(* Logix 5000 project; controller PLC_MCC1300_75F1 vendor 1 type 14 code 166 rev 32.11; software revision 32.04; part 65 of 83 *)
(* tags used below, declared in another part *)
   CM_AreaStackerToLine_JS1 : CM_AreaStackerToLine;
   CM_AreaStackerToLine_JS1_Sync : CM_AreaStackerToLine;
   CONST_dDest_Cullet : DINT;
   CONST_dDest_Stk : DINT;
   CONST_rgdDestMask : DINT[32];   // Destination Mask
   Convoy_SL_DATA_NULL : UDT_Convoy_SL;
   GP_AccessArea_M316S_STC : GP_AccessArea_STC;
   GP_CheckIdPlatePresent : GP_CheckIdPlatePresent;
   GP_InvertCapxLite : GP_InvertCapxLite;
   GP_M316A : GP_Rotator;
   GP_OB_InitializeMain : GP_OB_Initialize;
   GP_RampSpace : GP_RampSpace;
   Gp_SpaceConvUtilities_V1 : GP_SpaceConvUtilities_V1;
   M310B : MAC_Conveyor;
   M310B_Data : UDT_Convoy_SL;
   M310B_SpaceConv_Utilities : SpaceConv_Utilities;
   M312 : MAC_Conveyor_Single;
   M312_SpaceConv_Utilities : SpaceConv_Utilities;
   M315A_SpaceConv_Utilities : SpaceConv_Utilities;
   M315B : MAC_Conveyor;
   M315B_Data : UDT_Convoy_SL;
   M315B_SpaceConv_Utilities : SpaceConv_Utilities;
   M316 : MAC_Conveyor;
   M316_ALM : MAC_Conveyor_ALM;
   M316_Data : UDT_Convoy_SL;
   M316_dLastRotationA_ID : DINT;
   M316_HMW : MAC_Conveyor_HMW;
   M316_M1_DR_IN_MAM : MOTION_INSTRUCTION;
   M316_SpaceConv_Utilities : SpaceConv_Utilities;
   M316_xOS_SentToCullet : BOOL;
   M316_xPlateCullet : BOOL;
   M316_xSendCulletReqActive : BOOL;
   M316A : MAC_Rotator;
   M316A_Data : UDT_Convoy_SL;
   M316A_HMR : MAC_Rotator_HMR;
   M316A_HMW : MAC_Rotator_HMW;
   M316A_M1_DR : AXIS_CIP_DRIVE;
   M316A_M1_DR_IN_MAM : MOTION_INSTRUCTION;
   M316A_rLastPosition : REAL;
   M317_SpaceConv_Utilities : SpaceConv_Utilities;
   Sbr_OUT_ReqRot_CW : BOOL;
   TMP_d : DINT;
   TMP_dActualOnLHS : DINT;
   TMP_dConveyorNumberForZoneCleaning : DINT;
   TMP_dDecelerationPositionEndConveyor : DINT;
   TMP_dMissingOnLHS : DINT;
   TMP_dOffsetLoadUnload_cmm : DINT;
   TMP_dPhEndPosition_cmm : DINT;
   TMP_HeadPos : DINT;
   TMP_Portrait : BOOL;
   TMP_rgxId : DINT[10];
   TMP_x : BOOL;
   TMP_xConveyorInvolvedInCleaning : BOOL;
   TMP_xConveyorOfStartCleaning : BOOL;
   TMP_xCulletPresent : BOOL;
   TMP_xEnableLoadUnload : BOOL;
   TMP_xEnableZoneCleaning : BOOL;
   TMP_xJustOnePlateMissing : BOOL;
   TMP_xLiteThisDestPresent : BOOL;
   x316PortraitMode : BOOL;
   xAlwaysOFF : BOOL;
   xAlwaysON : BOOL;
   xDebugOFF : BOOL;
   Z402 : MAC_Zone;
   Z402_HMR : MAC_Zone_HMR;
   Z402_HMW : MAC_Zone_HMW;
(* MainProgram, continued *)

ROUTINE M316_Alarm   (* ladder *)
   // Reset Alarm
   0: XIC(Z402.tmON_ResetAlarm.DN)FLL(0,M316_ALM,1);
   1: XIC(Z402.ST_xEnableControlError)XIC(M316.INPUT_xDriveError_M1)OTL(M316_ALM.rgxStoppingFault_M[0].1);
   2: XIC(Z402.ST_xEnableControlError)XIO(M316.INPUT_xDriveError_M1)[XIC(M316.OUTPUT_xRun_M1) ,XIC(M316.OUTPUT_xReverse_M1) ,XIC(M316.OUTPUT_xPositioning_M1) ]XIO(M316.INPUT_xDriveFeedback_M1)[XIO(M316.tmON_FeedbackTimeOut_M1.DN) TON(M316.tmON_FeedbackTimeOut_M1,?,?) ,XIC(M316.tmON_FeedbackTimeOut_M1.DN) OTL(M316_ALM.rgxStoppingFault_M[0].2) ];
   3: XIC(Z402.ST_xEnableControlError)XIO(M316.INPUT_xMotorThermalProbe_M1)OTL(M316_ALM.rgxStoppingFault_M[0].4);
   4: XIC(Z402.ST_xEnableControlError)[XIC(M316.INPUT_xDriveInhibit_M1) ,XIC(M316.OUTPUT_xDriveEnable_M1) XIO(M316.INPUT_xDriveReady_M1) ][XIO(M316.tmON_DriveInhibit_M1.DN) TON(M316.tmON_DriveInhibit_M1,?,?) ,XIC(M316.tmON_DriveInhibit_M1.DN) OTL(M316_ALM.rgxStoppingFault_M[0].6) ];
   5: XIC(Z402.ST_xEnableControlError)XIC(M316.INPUT_xDriveError_M2)OTL(M316_ALM.rgxStoppingFault_M[0].11);
   6: XIC(Z402.ST_xEnableControlError)XIO(M316.INPUT_xDriveError_M2)[XIC(M316.OUTPUT_xRun_M2) ,XIC(M316.OUTPUT_xReverse_M2) ,XIC(M316.OUTPUT_xPositioning_M2) ]XIO(M316.INPUT_xDriveFeedback_M2)[XIO(M316.tmON_FeedbackTimeOut_M2.DN) TON(M316.tmON_FeedbackTimeOut_M2,?,?) ,XIC(M316.tmON_FeedbackTimeOut_M2.DN) OTL(M316_ALM.rgxStoppingFault_M[0].12) ];
   7: XIC(Z402.ST_xEnableControlError)XIO(M316.INPUT_xMotorThermalProbe_M2)OTL(M316_ALM.rgxStoppingFault_M[0].14);
   8: XIC(Z402.ST_xEnableControlError)[XIC(M316.INPUT_xDriveInhibit_M2) ,XIC(M316.OUTPUT_xDriveEnable_M2) XIO(M316.INPUT_xDriveReady_M2) ][XIO(M316.tmON_DriveInhibit_M2.DN) TON(M316.tmON_DriveInhibit_M2,?,?) ,XIC(M316.tmON_DriveInhibit_M2.DN) OTL(M316_ALM.rgxStoppingFault_M[0].16) ];
   9: XIC(M316.ST_xEnableControlError)XIC(M316.PH_x.7)NEQ(M316_SpaceConv_Utilities.CONST_dSyncMode,0)[XIO(M316.ST_xPlateSynchronized) OTL(M316_ALM.rgxWarning[0].0) ,XIC(M316.ST_xPlateSynchronized) OTU(M316_ALM.rgxWarning[0].0) ];
   10: XIC(M316.ST_xEnableControlError)[XIC(M316_Data.tFlag.tConveyor.xReqStop) [XIC(M316.PH_x.0) ,XIC(M316.PH_x.1) ] ADD(M316_SpaceConv_Utilities.CONST_dConveyorLength_cmm,200000,TMP_d) GRT(M316_SpaceConv_Utilities.O_dHeadPosition_cmm,TMP_d) ,XIC(M316.PH_x.16) CPT(TMP_d,M316_SpaceConv_Utilities.CONST_dConveyorLength_cmm + M316.AUX_dDecSpace_cmm) GRT(M316_SpaceConv_Utilities.O_dHeadPosition_cmm,TMP_d) ][OTL(M316_ALM.rgxWarning[0].1) ,OTL(M316.ST_xPhaseError) ];
   11: XIC(M316.ST_xEnableControlError)[XIC(M316.PH_x.0) ,XIC(M316.PH_x.8) ,XIC(M316.PH_x.16) ]XIO(M316A.INPUT_xLowPosition)OTL(M316_ALM.rgxStoppingFault[0].0);
   // #####_CUMULATIVE ALARM_#####
   12: NOP();
   13: [NEQ(M316_ALM.rgxStoppingFault[0],0) ,NEQ(M316_ALM.rgxStoppingFault_M[0],0) ,NEQ(M316_ALM.rgxStoppingFault_M[1],0) ]OTE(M316.ST_xStopMachineFault);
   14: [NEQ(M316_ALM.rgxFault[0],0) ,NEQ(M316_ALM.rgxFault_M[0],0) ,NEQ(M316_ALM.rgxFault_M[1],0) ]OTE(M316.ST_xStopNextCycleFault);
END_ROUTINE

ROUTINE M316_Logic   (* ladder *)
   // #####_COSTANTS_#####
   0: [MOV(4030,TMP_dConveyorNumberForZoneCleaning) MOV(350000,TMP_dOffsetLoadUnload_cmm) MOV(500,M316_SpaceConv_Utilities.CONST_dPresetFeedbackTime_ms) OTL(TMP_xEnableLoadUnload) OTU(TMP_xEnableZoneCleaning) MOV(450000,M316_SpaceConv_Utilities.CONST_dConveyorLength_cmm) MOV(375000,M316_SpaceConv_Utilities.CONST_dConveyorWidth_cmm) SUB(M316_SpaceConv_Utilities.CONST_dConveyorLength_cmm,M316.AUX_dAccSpace_cmm,M316.AUX_dPresetStopLoad_cmm) ADD(M316_SpaceConv_Utilities.CONST_dConveyorLength_cmm,M316.AUX_dDecSpace_cmm,M316.AUX_dPresetStopUnload_cmm) MOV(1.2,M316_SpaceConv_Utilities.CONST_rAcceleration_ms2) MOV(1.2,M316_SpaceConv_Utilities.CONST_rDeceleration_ms2) MOV(M316_SpaceConv_Utilities.CONST_dConveyorLength_cmm,TMP_dPhEndPosition_cmm) ,XIO(M316.PH_x.22) [MOV(1,M316_SpaceConv_Utilities.CONST_dSyncMode) ,MOV(25000,M316_SpaceConv_Utilities.CONST_dSyncroPhPosition_cmm) ,MOV(200000,M316_SpaceConv_Utilities.CONST_dSyncroPhWindow_cmm) ] ,XIC(M316.PH_x.22) [MOV(1,M316_SpaceConv_Utilities.CONST_dSyncMode) ,MOV(0,M316_SpaceConv_Utilities.CONST_dSyncroPhPosition_cmm) ,MOV(300000,M316_SpaceConv_Utilities.CONST_dSyncroPhWindow_cmm) ] ];
   // #####_MATCH_#####
   1: NOP();
   // Conveyor Cleaning
   2: XIC(TMP_xEnableZoneCleaning)XIC(Z402.ST_xCleaningAccepted)GRT(Z402_HMW.dCleaningSelection,0)[EQU(Z402_HMW.dCleaningSelection,TMP_dConveyorNumberForZoneCleaning) OTE(TMP_xConveyorOfStartCleaning) ,GEQ(Z402_HMW.dCleaningSelection,TMP_dConveyorNumberForZoneCleaning) OTE(TMP_xConveyorInvolvedInCleaning) ];
   // Enable control error
   3: XIC(Z402.ST_xEnableControlError)OTE(M316.ST_xEnableControlError);
   // Mode 7 - Offsett for load/unload Simultaney
   4: XIC(M316.PH_x.8)MOV(M316.AUX_dPresetStopLoad_cmm,M316_SpaceConv_Utilities.ST_dStopLoadForseen_cmm)MOV(TMP_dOffsetLoadUnload_cmm,M316_SpaceConv_Utilities.CONF_MD7_dOffset_cmm)GP_SpaceConvUtilities_V1(Gp_SpaceConvUtilities_V1,M316_SpaceConv_Utilities,M315A_SpaceConv_Utilities,M317_SpaceConv_Utilities,7);
   // #####_ALARMS_#####
   5: NOP();
   // Call Alarm Routine
   6: JSR(M316_Alarm,0);
   // Call Alarm Routine
   7: JSR(M316A_Rotator_Alarm,0);
   // #####_HMI_LOGICS_#####
   8: NOP();
   // Condition ok for Cleaning
   9: [XIO(TMP_xEnableZoneCleaning) ,XIC(TMP_xEnableZoneCleaning) XIC(M316.ST_xOutputEnable) [XIO(TMP_xConveyorOfStartCleaning) ,XIC(M316.PH_x.0) ,XIO(M316.PH_x.8) ] ]OTE(M316.ST_xCleaningConditionOK);
   // Cleaning Accepted
   10: [[XIC(M316_HMW.xStopLocalCleaningRequest) ,XIC(Z402_HMW.xStopCleanZoneRequest) ] OTU(M316_HMW.xStopLocalCleaningRequest) OTU(M316_HMW.xLocalCleaningRequest) ,[XIC(M316_HMW.xLocalCleaningRequest) ,XIC(xAlwaysOFF) XIC(M316.ST_xCleaningAccepted) XIC(TMP_xEnableZoneCleaning) ,XIO(xAlwaysOFF) XIC(Z402.ST_xCleaningAccepted) ] [XIC(M316.ST_xCleaningConditionOK) ,XIC(M316.ST_xCleaningAccepted) ] OTE(M316.ST_xCleaningAccepted) ];
   // Manual Mode Enabled
   11: XIO(M316_SpaceConv_Utilities.ST_xFeedbackRotation)[XIC(M316_HMW.xEnableDisableManualCommand) XIC(M316.ST_xConditionOKStopCycle) OTL(M316.ST_xManualMode) ,XIO(M316_HMW.xEnableDisableManualCommand) OTU(M316.ST_xManualMode) ];
   // Virtual door enabled
   12: XIC(M316_HMW.xEnableDisableVirtualDoor)OTE(M316.ST_xVirtualDoorEnabled);
   // Clear manual command
   13: [XIO(M316.ST_xManualMode) MOV(0,M316_HMW.rgxMan) ,XIO(M316A.ST_xManualMode) MOV(0,M316A_HMW.rgxMan) ];
   // #####_STATUSES_#####
   14: NOP();
   // Syncro  -  OS Syncro Photocell
   15: XIC(xAlwaysON)[[XIO(M316.PH_x.22) [XIC(M316.INPUT_xSyncroPhotocell_1) ,XIC(M316.PH_x.0) XIC(M316.INPUT_xSyncroPhotocell_2) ] ,XIC(xAlwaysOFF) XIC(M316.PH_x.22) XIC(M312.INPUT_xSyncroPhotocell_1) ] ONS(M316.OSR_xSynchroPhotocellHead) OTE(M316.OS_xSynchroPhotocellHead) GEQ(M316_SpaceConv_Utilities.CONST_dSyncMode,1) OTE(M316_SpaceConv_Utilities.ST_OS_xSynchroPhotocellHead) ,[XIO(M316.PH_x.22) XIO(M316.INPUT_xSyncroPhotocell_1) XIO(M316.INPUT_xSyncroPhotocell_2) ,XIC(xAlwaysOFF) XIC(M316.PH_x.22) XIO(M312.INPUT_xSyncroPhotocell_1) ] ONS(M316.OSR_xSynchroPhotocellTail) OTE(M316.OS_xSynchroPhotocellTail) GEQ(M316_SpaceConv_Utilities.CONST_dSyncMode,2) OTE(M316_SpaceConv_Utilities.ST_OS_xSynchroPhotocellTail) ];
   // Id Plate presence
   16: MOV(CONST_rgdDestMask[24],CONST_dDest_Cullet)GP_CheckIdPlatePresent(GP_CheckIdPlatePresent,M316_Data,TMP_rgxId,M316.ST_xIdPlatePresence,TMP_xCulletPresent,CONST_dDest_Cullet)MOV(CONST_rgdDestMask[1],CONST_dDest_Stk)GP_CheckIdPlatePresent(GP_CheckIdPlatePresent,M316_Data,TMP_rgxId,M316.ST_xIdPlatePresence,TMP_xLiteThisDestPresent,CONST_dDest_Stk)XIC(TMP_xCulletPresent)OTE(M316_xPlateCullet);
   // Machine in Alarm
   17: [XIC(M316.ST_xStopMachineFault) ,XIC(M316.ST_xStopNextCycleFault) ]OTE(M316.ST_xMachineAlarm);
   // Condition ok for stop Cycle
   18: [XIO(M316.ST_xPhasesInProgress) ,XIC(M316.PH_x.8) XIO(M316.OUTPUT_xRun_M1) XIO(M316_SpaceConv_Utilities.ST_xFeedbackRotation) XIO(M316.OUTPUT_xRun_M2) ,XIC(M316.ST_xMachineAlarm) ,XIO(Z402.ST_xCycleON) ]OTE(M316.ST_xConditionOKStopCycle);
   // Cycle load unload simultaneous
   19: XIC(TMP_xEnableLoadUnload)XIO(M316.ST_xDisableLoadUnloadOnStop)XIO(M316.ST_xIdPlatePresence)OTE(M316.ST_xCycleLoadUnload);
   // Speed Management
   20: [XIO(M316_SpaceConv_Utilities.O_xRampInProgress) XIO(M316.ST_xManualMode) MOV(Z402_HMR.dLineSpeed_mm_min,M316.AUX_dReqSpeed_mm_min) ,XIC(M316.ST_xManualMode) MOV(Z402_HMW.dManualSpeed_mm_min,M316.AUX_dReqSpeed_mm_min) ,NEQ(M316.AUX_dReqSpeed_mm_min,M316_SpaceConv_Utilities.ST_dRealSpeed_mm_min) OTE(M316.OS_xChangeSpeed) ];
   // Ramp Management
   21: GP_RampSpace(GP_RampSpace,M316_SpaceConv_Utilities.CONST_rAcceleration_ms2,M316_SpaceConv_Utilities.CONST_rDeceleration_ms2,M316_SpaceConv_Utilities.ST_dRealSpeed_mm_min,M316.AUX_dAccSpace_cmm,M316.AUX_dDecSpace_cmm);
   // Space Convoy utilities MOD 1 for Calculate Head/Tail
   22: XIC(xAlwaysON)[[XIC(M316.OUTPUT_xRun_M1) ,XIC(M316.OUTPUT_xReverse_M1) ] XIO(M316.ST_xManualMode) OTE(M316_SpaceConv_Utilities.CONF_MD1_xRun) ,XIC(M316.OUTPUT_xReverse_M1) XIC(xAlwaysOFF) XIO(M316.ST_xManualMode) OTE(M316_SpaceConv_Utilities.CONF_MD1_xReverse) ,[XIC(M316.INPUT_xDriveFeedback_M1) ,XIC(M316_SpaceConv_Utilities.CONF_MD1_xRun) GRT(M316_SpaceConv_Utilities.O_dCountFeedbackTime_ms,0) ] OTE(M316_SpaceConv_Utilities.ST_xFeedbackRotation) ,XIC(M316.ST_xIdPlatePresence) OTE(M316_SpaceConv_Utilities.CONF_MD1_xHeadTracking) ,XIC(M316.ST_xPlatePresence) OTE(M316_SpaceConv_Utilities.CONF_MD1_xTailTracking) ,MOV(GP_OB_InitializeMain.OUT_dExecutionTime_ms,M316_SpaceConv_Utilities.CONF_MD1_dScan_ms) GP_SpaceConvUtilities_V1(Gp_SpaceConvUtilities_V1,M316_SpaceConv_Utilities,M315A_SpaceConv_Utilities,M317_SpaceConv_Utilities,1) ];
   // Output Enable
   23: XIC(Z402.ST_xCycleON)XIO(M316.ST_xManualMode)XIO(M316.ST_xStopMachineFault)[XIO(M316.ST_xPlatePassageUpstream_FW) XIO(M316.ST_xPlatePassageUpstream_BKW) ,XIC(M316.ST_xPlatePassageUpstream_FW) XIC(M310B.ST_xOutputEnable) ,XIC(M316.ST_xPlatePassageUpstream_BKW) XIC(M312.ST_xOutputEnable) ]XIC(M316A.INPUT_xLowPosition)OTE(M316.ST_xOutputEnable);
   24: XIO(TMP_xLiteThisDestPresent)OTU(M316_xSendCulletReqActive);
   // #####_WORKING_FLAGS_#####
   25: NOP();
   // #####_LOGICS_#####
   26: NOP();
   // Phase of load
   27: XIC(M310B.OS_xUnload_FW)[[XIC(M310B.PH_x.8) ,XIC(M310B.PH_x.16) ] OTL(M316.PH_x.0) ,OTU(M316_SpaceConv_Utilities.O_xPlateSynchronized) ,OTU(M316.ST_xDisableLoadUnloadOnStop) ,OTE(M316.OS_xLoad_FW) ,XIC(M315B.OS_xUnload_FW) COP(M310B_Data,M316_Data,1) FLL(0,M310B_Data,1) ,GP_SpaceConvUtilities_V1(Gp_SpaceConvUtilities_V1,M316_SpaceConv_Utilities,M315A_SpaceConv_Utilities,M317_SpaceConv_Utilities,5) ,XIC(M315B.OS_xUnpack) ADD(M310B_SpaceConv_Utilities.O_dTailPosition_cmm,M315B_Data.dLength_cmm,M315B_SpaceConv_Utilities.CONF_MD2_MD3_dPrstPos_cmm) GP_SpaceConvUtilities_V1(Gp_SpaceConvUtilities_V1,M315B_SpaceConv_Utilities,M315B_SpaceConv_Utilities,M315A_SpaceConv_Utilities,2) ];
   // Request Rotation
   // Inserire le condizioni per far ruotare le lastre (stacker, lastre in arrivo etc)
   28: [[XIC(M310B.OS_xUnload_FW) ,XIC(M310B.OS_xUnpack) ] [NEQ(M316_Data.rgtCap[0].rgtLite[0].dID,0) GRT(M316_Data.rgtCap[0].dLength_cmm,M316_Data.rgtCap[0].rgtLite[0].dWidth_cmm) OTE(TMP_Portrait) ,[XIC(TMP_Portrait) XIO(x316PortraitMode) ,XIO(TMP_Portrait) XIC(x316PortraitMode) [XIC(CM_AreaStackerToLine_JS1_Sync.xStackerInUnloaderMode) ,XIO(xAlwaysOFF) ] ] [LEQ(M316_Data.rgtCap[0].dNumLites,2) ,XIO(xAlwaysOFF) ] OTE(Sbr_OUT_ReqRot_CW) ] ,XIC(Sbr_OUT_ReqRot_CW) [XIC(xAlwaysON) OTL(M316_Data.tFlag.tRotator.xReqRotationCw) OTU(M316_Data.tFlag.tRotator.xReqRotationCcw) ,XIC(xAlwaysOFF) OTL(M316_Data.tFlag.tRotator.xReqRotationCcw) OTU(M316_Data.tFlag.tRotator.xReqRotationCw) ] ];
   // Request positioning
   29: [XIC(M310B.OS_xUnload_FW) ,XIC(M310B.OS_xUnpack) ][XIC(M316_Data.tFlag.tRotator.xReqRotationCw) ,XIC(M316_Data.tFlag.tRotator.xReqRotationCcw) ][OTL(M316_Data.tFlag.tConveyor.xReqStop) ,CPT(M316.AUX_dPhPosTarget_cmm,M316_SpaceConv_Utilities.CONST_dConveyorLength_cmm / 2 + M316_Data.dLength_cmm / 2 - M316_SpaceConv_Utilities.CONST_dSyncroPhPosition_cmm + M316_HMW.dParam_1_cmm + 5000) ];
   // Syncro  -  Space Convoy utilities MOD 4
   30: GRT(M316_SpaceConv_Utilities.CONST_dSyncMode,0)[XIC(M316.PH_x.0) XIO(M316.PH_x.8) ,XIC(M316.PH_x.0) XIC(M316.PH_x.8) ADD(M316_SpaceConv_Utilities.CONST_dSyncroPhPosition_cmm,TMP_dOffsetLoadUnload_cmm,TMP_d) GRT(M316_SpaceConv_Utilities.O_dTailPosition_cmm,TMP_d) ][MOV(M316_Data.dLength_cmm,M316_SpaceConv_Utilities.CONF_MD4_MD6_dLength_cmm) ,GP_SpaceConvUtilities_V1(Gp_SpaceConvUtilities_V1,M316_SpaceConv_Utilities,M315A_SpaceConv_Utilities,M317_SpaceConv_Utilities,4) ];
   // End load Phase
   31: XIC(M316.PH_x.0)[XIO(M316_Data.tFlag.tConveyor.xReqStop) GRT(M316_SpaceConv_Utilities.O_dHeadPosition_cmm,M316.AUX_dPresetStopLoad_cmm) ,XIC(M316_Data.tFlag.tConveyor.xReqStop) [XIC(M316.OUTPUT_xPositioning_M1) XIC(M316_M1_DR_IN_MAM.PC) ,XIC(M316.ST_xPhaseError) ] ][OTU(M316.PH_x.0) ,OTE(M316.PH_x.7) ,OTL(M316.ST_xPlatePresence) ];
   // End positiong
   32: XIC(M316.PH_x.7)XIC(M316_Data.tFlag.tConveyor.xReqStop)XIC(M316.OUTPUT_xPositioning_M1)XIC(M316_M1_DR_IN_MAM.PC)XIC(M316.OUTPUT_xPositioning_M2)[OTU(M316_Data.tFlag.tConveyor.xReqStop) ,OTL(M316_Data.tFlag.tConveyor.xReqStopEndConveyor) ,CPT(M316_SpaceConv_Utilities.CONF_MD2_MD3_dPrstPos_cmm,M316.AUX_dPhPosTarget_cmm + M316_SpaceConv_Utilities.CONST_dSyncroPhPosition_cmm - M316_HMW.dParam_1_cmm) GP_SpaceConvUtilities_V1(Gp_SpaceConvUtilities_V1,M316_SpaceConv_Utilities,M315A_SpaceConv_Utilities,M316_SpaceConv_Utilities,2) XIC(xAlwaysOFF) GP_SpaceConvUtilities_V1(Gp_SpaceConvUtilities_V1,M316_SpaceConv_Utilities,M315A_SpaceConv_Utilities,M317_SpaceConv_Utilities,2) ];
   // Calculation Space for Wait Stop Next Conveyor
   33: CPT(TMP_dDecelerationPositionEndConveyor,M316_SpaceConv_Utilities.CONST_dConveyorLength_cmm - M316.AUX_dAccSpace_cmm + 1000);
   // Wait stop next Machine
   34: XIO(M316.PH_x.8)GEQ(M316_SpaceConv_Utilities.O_dHeadPosition_cmm,TMP_dDecelerationPositionEndConveyor)OTE(M316.ST_xWaitStopNextMachine);
   // Set Wait Machine Stop
   35: [XIC(M316.PH_x.7) [XIO(M312.ST_xInitialConditionOK) ,XIC(M316.ST_xWaitStopNextMachine) [XIC(M312_SpaceConv_Utilities.O_xRampInProgress) ,XIO(M312_SpaceConv_Utilities.ST_xFeedbackRotation) ] ] ,XIC(M316.PH_x.0) NEQ(Z402_HMR.dLineSpeed_mm_min,M316.AUX_dReqSpeed_mm_min) ]OTL(M316.ST_xWaitMachineStop);
   // Reset Wait Machine Stop
   36: XIO(M316_SpaceConv_Utilities.ST_xFeedbackRotation)[XIO(M316_SpaceConv_Utilities.ST_xFeedbackRotation) ,XIO(M316.ST_xWaitStopNextMachine) ]EQU(Z402_HMR.dLineSpeed_mm_min,M316.AUX_dReqSpeed_mm_min)OTU(M316.ST_xWaitMachineStop);
   37: XIC(Z402.ST_xConditionOkPhaseAdvancement)XIC(M316.ST_xOutputEnable)XIC(M316.ST_xPlatePresence)XIC(M316.ST_xIdPlatePresence)XIO(M316.ST_xWaitMachineStop)XIO(M316.ST_xPhasesInProgress)OTE(M316.ST_xWaitReadyToMove);
   38: XIO(xDebugOFF)MOV(0,TMP_dActualOnLHS);
   39: SUB(CM_AreaStackerToLine_JS1.iPresetNumberPlateOnRack[0],TMP_dActualOnLHS,TMP_dMissingOnLHS)EQU(TMP_dMissingOnLHS,1)[EQU(CM_AreaStackerToLine_JS1.iActualNumberPlateOnRack[0],0) ,EQU(CM_AreaStackerToLine_JS1.iActualNumberPlateOnRack[0],CM_AreaStackerToLine_JS1.iPresetNumberPlateOnRack[0]) ]OTE(TMP_xJustOnePlateMissing);
   // Phase of unload
   40: XIO(M316_xSendCulletReqActive)XIC(Z402.ST_xConditionOkPhaseAdvancement)XIC(M316.ST_xPlatePresence)XIC(M316.ST_xIdPlatePresence)XIC(M316.ST_xOutputEnable)XIC(M312.ST_xInitialConditionOK)XIO(M316.ST_xWaitMachineStop)XIO(M316.PH_x.8)[XIO(M316_Data.tFlag.tRotator.xReqRotationCw) ,XIC(M316_Data.tFlag.tRotator.xDoneRotationCw) ][XIO(M316_Data.tFlag.tRotator.xReqRotationCcw) ,XIC(M316_Data.tFlag.tRotator.xDoneRotationCcw) ]XIC(TMP_xLiteThisDestPresent)XIO(M316.PH_x.8)[OTL(M316.PH_x.8) ,OTE(M316.OS_xUnload_FW) ,MOV(M316_Data.dLength_cmm,M316_SpaceConv_Utilities.CONF_MD4_MD6_dLength_cmm) GP_SpaceConvUtilities_V1(Gp_SpaceConvUtilities_V1,M316_SpaceConv_Utilities,M315A_SpaceConv_Utilities,M317_SpaceConv_Utilities,6) ];
   // Phase of end unload
   41: XIC(M316.PH_x.8)[GEQ(M316_SpaceConv_Utilities.O_dTailPosition_cmm,M316.AUX_dPresetStopUnload_cmm) ,XIO(M316_SpaceConv_Utilities.ST_xFeedbackRotation) GEQ(M316_SpaceConv_Utilities.O_dTailPosition_cmm,M316_SpaceConv_Utilities.CONST_dConveyorLength_cmm) ][OTE(M316.PH_x.15) ,OTU(M316.PH_x.8) ,OTU(M316.ST_xPlatePresence) ];
   // Rotator managment
   // -
   // -
   42: NOP();
   43: XIO(M316_xSendCulletReqActive)XIC(M316.ST_xPlatePresence)XIC(M316.ST_xIdPlatePresence)XIO(M316.ST_xPhasesInProgress)XIO(M316.ST_xStopMachineFault)[XIC(M316_Data.tFlag.tRotator.xReqRotationCw) ,XIC(M316_Data.tFlag.tRotator.xReqRotationCcw) ]XIO(M316_Data.tFlag.tConveyor.xReqStop)XIO(M316_Data.tFlag.tConveyor.xBypassReqEndStop)XIC(M316_Data.tFlag.tConveyor.xReqStopEndConveyor)NEQ(M316_Data.rgtCap[0].rgtLite[0].dID,M316_dLastRotationA_ID)COP(M316_Data,M316A_Data,1)[OTL(M316.PH_x.3) ,MOV(M316_Data.rgtCap[0].rgtLite[0].dID,M316_dLastRotationA_ID) ,MOV(M316A_M1_DR.ActualPosition,M316A_rLastPosition) ];
   44: [XIC(GP_AccessArea_M316S_STC.ST_xAccessRequest) OTE(GP_M316A.IN_xReqAccess) ,XIC(xDebugOFF) OTE(GP_M316A.IN_xDoneAccess) ,XIC(M316A.INPUT_xConditionToDescent) OTE(GP_M316A.IN_xConditionToDescent) ,XIC(M316A.INPUT_xDriveFeedback) OTE(GP_M316A.IN_xDriveFeedback) ,XIC(M316A.INPUT_xHighPosition) OTE(GP_M316A.IN_xHighPosition) ,XIC(M316A.INPUT_xLowPosition) OTE(GP_M316A.IN_xLowPosition) ,[XIC(M316A_M1_DR_IN_MAM.EN) ,XIO(xAlwaysOFF) ] [XIC(M316A_M1_DR_IN_MAM.PC) ,XIO(xAlwaysOFF) [GEQ(M316A_rLastPosition,359.8) LEQ(M316A_rLastPosition,0.2) GEQ(M316A_M1_DR.ActualPosition,89.8) LEQ(M316A_M1_DR.ActualPosition,90.2) ,GEQ(M316A_rLastPosition,89.8) LEQ(M316A_rLastPosition,90.2) GEQ(M316A_M1_DR.ActualPosition,179.8) LEQ(M316A_M1_DR.ActualPosition,180.2) ,GEQ(M316A_rLastPosition,179.8) LEQ(M316A_rLastPosition,180.2) GEQ(M316A_M1_DR.ActualPosition,269.8) LEQ(M316A_M1_DR.ActualPosition,270.2) ,GEQ(M316A_rLastPosition,269.8) LEQ(M316A_rLastPosition,270.2) GEQ(M316A_M1_DR.ActualPosition,359.8) LEQ(M316A_M1_DR.ActualPosition,0.2) ] ] OTE(GP_M316A.IN_xPositionReached) ,XIC(Z402.ST_xCycleON) OTE(TMP_x) ,MOV(0,GP_M316A.IN_dWander_cmm) ,MOV(M316A.INPUT_rRotatorPosition_cdeg,GP_M316A.IN_dRotatorPosition_cdeg) ,GP_Rotator(GP_M316A,M316A,M316A_HMR,M316A_HMW,M316A_Data,TMP_x,Z402.ST_xConditionOkPhaseAdvancement,M316.ST_xManualMode,M316A_Data.tFlag.tRotator,TMP_HeadPos) ,XIC(M316A.INPUT_xLowPosition) OTE(M316A_HMR.xLowPosition) ];
   45: XIC(M316.PH_x.3)[XIC(M316A_Data.tFlag.tRotator.xDoneRotationCw) ,XIC(M316A_Data.tFlag.tRotator.xDoneRotationCcw) ]XIC(M316A.INPUT_xLowPosition)[OTE(M316.PH_x.4) ,OTU(M316.PH_x.3) ];
   46: XIC(M316.PH_x.4)[[XIC(M316A_Data.tFlag.tRotator.xDoneRotationCw) MOV(2,GP_InvertCapxLite.In_dOutDirection) ,XIC(M316A_Data.tFlag.tRotator.xDoneRotationCcw) MOV(3,GP_InvertCapxLite.In_dOutDirection) ] DIV(M316_SpaceConv_Utilities.CONST_dConveyorLength_cmm,2,GP_InvertCapxLite.In_dOffset1) GP_InvertCapxLite(GP_InvertCapxLite,1,1,GP_InvertCapxLite.In_dOutDirection,M316A_Data,M316_Data,Convoy_SL_DATA_NULL,M316_SpaceConv_Utilities.CONST_dConveyorLength_cmm,M316_SpaceConv_Utilities.CONST_dConveyorWidth_cmm,M316_SpaceConv_Utilities.CONF_MD2_MD3_dPrstPos_cmm,M316_SpaceConv_Utilities.O_dHeadPosition_cmm,GP_InvertCapxLite.In_dOffset1) [NEQ(M316A_Data.rgtCap[0].dID,0) MOV(M316A_Data.rgtCap[0].dThickness_cmm,M316_Data.rgtCap[0].dThickness_cmm) ,FLL(0,M316A_Data,1) ] ,CPT(M316_Data.dGapCaps_cmm,M316_Data.dLength_cmm-M316_Data.rgtCap[0].dLength_cmm-M316_Data.rgtCap[1].dLength_cmm) MOV(TMP_HeadPos,M316_SpaceConv_Utilities.O_dHeadPosition_cmm) ];
   47: XIC(M316.ST_xPhaseError)XIC(M316_xOS_SentToCullet)OTU(M316.ST_xPhaseError);
